   "SDC_EMS01_Carrier74_Faulted" AT %Q10841.6 : Bool;
   "SDC_EMS01_Carrier74_InAuto" AT %Q10841.7 : Bool;
   "SDC_EMS01_Carrier75_Spare0" AT %Q10842.0 : Bool;
   "SDC_EMS01_Carrier75_DriveTripped" AT %Q10842.1 : Bool;
   "SDC_EMS01_Carrier75_Spare2" AT %Q10842.2 : Bool;
   "SDC_EMS01_Carrier75_PositioningComplete" AT %Q10842.3 : Bool;
   "SDC_EMS01_Carrier75_RunStopPressed" AT %Q10842.4 : Bool;
   "SDC_EMS01_Carrier75_Moving" AT %Q10842.5 : Bool;
   "SDC_EMS01_Carrier75_Faulted" AT %Q10842.6 : Bool;
   "SDC_EMS01_Carrier75_InAuto" AT %Q10842.7 : Bool;
   "SDC_EMS01_Carrier76_Spare0" AT %Q10843.0 : Bool;
   "SDC_EMS01_Carrier76_DriveTripped" AT %Q10843.1 : Bool;
   "SDC_EMS01_Carrier76_Spare2" AT %Q10843.2 : Bool;
   "SDC_EMS01_Carrier76_PositioningComplete" AT %Q10843.3 : Bool;
   "SDC_EMS01_Carrier76_RunStopPressed" AT %Q10843.4 : Bool;
   "SDC_EMS01_Carrier76_Moving" AT %Q10843.5 : Bool;
   "SDC_EMS01_Carrier76_Faulted" AT %Q10843.6 : Bool;
   "SDC_EMS01_Carrier76_InAuto" AT %Q10843.7 : Bool;
   "SDC_EMS01_Carrier77_Spare0" AT %Q10844.0 : Bool;
   "SDC_EMS01_Carrier77_DriveTripped" AT %Q10844.1 : Bool;
   "SDC_EMS01_Carrier77_Spare2" AT %Q10844.2 : Bool;
   "SDC_EMS01_Carrier77_PositioningComplete" AT %Q10844.3 : Bool;
   "SDC_EMS01_Carrier77_RunStopPressed" AT %Q10844.4 : Bool;
   "SDC_EMS01_Carrier77_Moving" AT %Q10844.5 : Bool;
   "SDC_EMS01_Carrier77_Faulted" AT %Q10844.6 : Bool;
   "SDC_EMS01_Carrier77_InAuto" AT %Q10844.7 : Bool;
   "SDC_EMS01_Carrier78_Spare0" AT %Q10845.0 : Bool;
   "SDC_EMS01_Carrier78_DriveTripped" AT %Q10845.1 : Bool;
   "SDC_EMS01_Carrier78_Spare2" AT %Q10845.2 : Bool;
   "SDC_EMS01_Carrier78_PositioningComplete" AT %Q10845.3 : Bool;
   "SDC_EMS01_Carrier78_RunStopPressed" AT %Q10845.4 : Bool;
   "SDC_EMS01_Carrier78_Moving" AT %Q10845.5 : Bool;
   "SDC_EMS01_Carrier78_Faulted" AT %Q10845.6 : Bool;
   "SDC_EMS01_Carrier78_InAuto" AT %Q10845.7 : Bool;
   "SDC_EMS01_Carrier79_Spare0" AT %Q10846.0 : Bool;
   "SDC_EMS01_Carrier79_DriveTripped" AT %Q10846.1 : Bool;
   "SDC_EMS01_Carrier79_Spare2" AT %Q10846.2 : Bool;
   "SDC_EMS01_Carrier79_PositioningComplete" AT %Q10846.3 : Bool;
   "SDC_EMS01_Carrier79_RunStopPressed" AT %Q10846.4 : Bool;
   "SDC_EMS01_Carrier79_Moving" AT %Q10846.5 : Bool;
   "SDC_EMS01_Carrier79_Faulted" AT %Q10846.6 : Bool;
   "SDC_EMS01_Carrier79_InAuto" AT %Q10846.7 : Bool;
   "SDC_EMS01_Carrier80_Spare0" AT %Q10847.0 : Bool;
   "SDC_EMS01_Carrier80_DriveTripped" AT %Q10847.1 : Bool;
   "SDC_EMS01_Carrier80_Spare2" AT %Q10847.2 : Bool;
   "SDC_EMS01_Carrier80_PositioningComplete" AT %Q10847.3 : Bool;
   "SDC_EMS01_Carrier80_RunStopPressed" AT %Q10847.4 : Bool;
   "SDC_EMS01_Carrier80_Moving" AT %Q10847.5 : Bool;
   "SDC_EMS01_Carrier80_Faulted" AT %Q10847.6 : Bool;
   "SDC_EMS01_Carrier80_InAuto" AT %Q10847.7 : Bool;
   "SDC_EMS01_Carrier81_Spare0" AT %Q10848.0 : Bool;
   "SDC_EMS01_Carrier81_DriveTripped" AT %Q10848.1 : Bool;
   "SDC_EMS01_Carrier81_Spare2" AT %Q10848.2 : Bool;
   "SDC_EMS01_Carrier81_PositioningComplete" AT %Q10848.3 : Bool;
   "SDC_EMS01_Carrier81_RunStopPressed" AT %Q10848.4 : Bool;
   "SDC_EMS01_Carrier81_Moving" AT %Q10848.5 : Bool;
   "SDC_EMS01_Carrier81_Faulted" AT %Q10848.6 : Bool;
   "SDC_EMS01_Carrier81_InAuto" AT %Q10848.7 : Bool;
   "SDC_EMS01_Carrier82_Spare0" AT %Q10849.0 : Bool;
   "SDC_EMS01_Carrier82_DriveTripped" AT %Q10849.1 : Bool;
   "SDC_EMS01_Carrier82_Spare2" AT %Q10849.2 : Bool;
   "SDC_EMS01_Carrier82_PositioningComplete" AT %Q10849.3 : Bool;
   "SDC_EMS01_Carrier82_RunStopPressed" AT %Q10849.4 : Bool;
   "SDC_EMS01_Carrier82_Moving" AT %Q10849.5 : Bool;
   "SDC_EMS01_Carrier82_Faulted" AT %Q10849.6 : Bool;
   "SDC_EMS01_Carrier82_InAuto" AT %Q10849.7 : Bool;
   "SDC_EMS01_Carrier83_Spare0" AT %Q10850.0 : Bool;
   "SDC_EMS01_Carrier83_DriveTripped" AT %Q10850.1 : Bool;
   "SDC_EMS01_Carrier83_Spare2" AT %Q10850.2 : Bool;
   "SDC_EMS01_Carrier83_PositioningComplete" AT %Q10850.3 : Bool;
   "SDC_EMS01_Carrier83_RunStopPressed" AT %Q10850.4 : Bool;
   "SDC_EMS01_Carrier83_Moving" AT %Q10850.5 : Bool;
   "SDC_EMS01_Carrier83_Faulted" AT %Q10850.6 : Bool;
   "SDC_EMS01_Carrier83_InAuto" AT %Q10850.7 : Bool;
   "SDC_EMS01_Carrier84_Spare0" AT %Q10851.0 : Bool;
   "SDC_EMS01_Carrier84_DriveTripped" AT %Q10851.1 : Bool;
   "SDC_EMS01_Carrier84_Spare2" AT %Q10851.2 : Bool;
   "SDC_EMS01_Carrier84_PositioningComplete" AT %Q10851.3 : Bool;
   "SDC_EMS01_Carrier84_RunStopPressed" AT %Q10851.4 : Bool;
   "SDC_EMS01_Carrier84_Moving" AT %Q10851.5 : Bool;
   "SDC_EMS01_Carrier84_Faulted" AT %Q10851.6 : Bool;
   "SDC_EMS01_Carrier84_InAuto" AT %Q10851.7 : Bool;
   "SDC_EMS01_Carrier85_Spare0" AT %Q10852.0 : Bool;
   "SDC_EMS01_Carrier85_DriveTripped" AT %Q10852.1 : Bool;
   "SDC_EMS01_Carrier85_Spare2" AT %Q10852.2 : Bool;
   "SDC_EMS01_Carrier85_PositioningComplete" AT %Q10852.3 : Bool;
   "SDC_EMS01_Carrier85_RunStopPressed" AT %Q10852.4 : Bool;
   "SDC_EMS01_Carrier85_Moving" AT %Q10852.5 : Bool;
   "SDC_EMS01_Carrier85_Faulted" AT %Q10852.6 : Bool;
   "SDC_EMS01_Carrier85_InAuto" AT %Q10852.7 : Bool;
   "SDC_EMS01_Carrier86_Spare0" AT %Q10853.0 : Bool;
   "SDC_EMS01_Carrier86_DriveTripped" AT %Q10853.1 : Bool;
   "SDC_EMS01_Carrier86_Spare2" AT %Q10853.2 : Bool;
   "SDC_EMS01_Carrier86_PositioningComplete" AT %Q10853.3 : Bool;
   "SDC_EMS01_Carrier86_RunStopPressed" AT %Q10853.4 : Bool;
   "SDC_EMS01_Carrier86_Moving" AT %Q10853.5 : Bool;
   "SDC_EMS01_Carrier86_Faulted" AT %Q10853.6 : Bool;
   "SDC_EMS01_Carrier86_InAuto" AT %Q10853.7 : Bool;
   "SDC_EMS01_Carrier87_Spare0" AT %Q10854.0 : Bool;
   "SDC_EMS01_Carrier87_DriveTripped" AT %Q10854.1 : Bool;
   "SDC_EMS01_Carrier87_Spare2" AT %Q10854.2 : Bool;
   "SDC_EMS01_Carrier87_PositioningComplete" AT %Q10854.3 : Bool;
   "SDC_EMS01_Carrier87_RunStopPressed" AT %Q10854.4 : Bool;
   "SDC_EMS01_Carrier87_Moving" AT %Q10854.5 : Bool;
   "SDC_EMS01_Carrier87_Faulted" AT %Q10854.6 : Bool;
   "SDC_EMS01_Carrier87_InAuto" AT %Q10854.7 : Bool;
   "SDC_EMS01_Carrier88_Spare0" AT %Q10855.0 : Bool;
   "SDC_EMS01_Carrier88_DriveTripped" AT %Q10855.1 : Bool;
   "SDC_EMS01_Carrier88_Spare2" AT %Q10855.2 : Bool;
   "SDC_EMS01_Carrier88_PositioningComplete" AT %Q10855.3 : Bool;
   "SDC_EMS01_Carrier88_RunStopPressed" AT %Q10855.4 : Bool;
   "SDC_EMS01_Carrier88_Moving" AT %Q10855.5 : Bool;
   "SDC_EMS01_Carrier88_Faulted" AT %Q10855.6 : Bool;
   "SDC_EMS01_Carrier88_InAuto" AT %Q10855.7 : Bool;
   "SDC_EMS01_Carrier89_Spare0" AT %Q10856.0 : Bool;
   "SDC_EMS01_Carrier89_DriveTripped" AT %Q10856.1 : Bool;
   "SDC_EMS01_Carrier89_Spare2" AT %Q10856.2 : Bool;
   "SDC_EMS01_Carrier89_PositioningComplete" AT %Q10856.3 : Bool;
   "SDC_EMS01_Carrier89_RunStopPressed" AT %Q10856.4 : Bool;
   "SDC_EMS01_Carrier89_Moving" AT %Q10856.5 : Bool;
   "SDC_EMS01_Carrier89_Faulted" AT %Q10856.6 : Bool;
   "SDC_EMS01_Carrier89_InAuto" AT %Q10856.7 : Bool;
   "SDC_EMS01_Carrier90_Spare0" AT %Q10857.0 : Bool;
   "SDC_EMS01_Carrier90_DriveTripped" AT %Q10857.1 : Bool;
   "SDC_EMS01_Carrier90_Spare2" AT %Q10857.2 : Bool;
   "SDC_EMS01_Carrier90_PositioningComplete" AT %Q10857.3 : Bool;
   "SDC_EMS01_Carrier90_RunStopPressed" AT %Q10857.4 : Bool;
   "SDC_EMS01_Carrier90_Moving" AT %Q10857.5 : Bool;
   "SDC_EMS01_Carrier90_Faulted" AT %Q10857.6 : Bool;
   "SDC_EMS01_Carrier90_InAuto" AT %Q10857.7 : Bool;
   "SDC_EMS01_Carrier91_Spare0" AT %Q10858.0 : Bool;
   "SDC_EMS01_Carrier91_DriveTripped" AT %Q10858.1 : Bool;
   "SDC_EMS01_Carrier91_Spare2" AT %Q10858.2 : Bool;
   "SDC_EMS01_Carrier91_PositioningComplete" AT %Q10858.3 : Bool;
   "SDC_EMS01_Carrier91_RunStopPressed" AT %Q10858.4 : Bool;
   "SDC_EMS01_Carrier91_Moving" AT %Q10858.5 : Bool;
   "SDC_EMS01_Carrier91_Faulted" AT %Q10858.6 : Bool;
   "SDC_EMS01_Carrier91_InAuto" AT %Q10858.7 : Bool;
   "SDC_EMS01_Carrier92_Spare0" AT %Q10859.0 : Bool;
   "SDC_EMS01_Carrier92_DriveTripped" AT %Q10859.1 : Bool;
   "SDC_EMS01_Carrier92_Spare2" AT %Q10859.2 : Bool;
   "SDC_EMS01_Carrier92_PositioningComplete" AT %Q10859.3 : Bool;
   "SDC_EMS01_Carrier92_RunStopPressed" AT %Q10859.4 : Bool;
   "SDC_EMS01_Carrier92_Moving" AT %Q10859.5 : Bool;
   "SDC_EMS01_Carrier92_Faulted" AT %Q10859.6 : Bool;
   "SDC_EMS01_Carrier92_InAuto" AT %Q10859.7 : Bool;
   "SDC_EMS01_Carrier93_Spare0" AT %Q10860.0 : Bool;
   "SDC_EMS01_Carrier93_DriveTripped" AT %Q10860.1 : Bool;
   "SDC_EMS01_Carrier93_Spare2" AT %Q10860.2 : Bool;
   "SDC_EMS01_Carrier93_PositioningComplete" AT %Q10860.3 : Bool;
   "SDC_EMS01_Carrier93_RunStopPressed" AT %Q10860.4 : Bool;
   "SDC_EMS01_Carrier93_Moving" AT %Q10860.5 : Bool;
   "SDC_EMS01_Carrier93_Faulted" AT %Q10860.6 : Bool;
   "SDC_EMS01_Carrier93_InAuto" AT %Q10860.7 : Bool;
   "SDC_EMS01_Carrier94_Spare0" AT %Q10861.0 : Bool;
   "SDC_EMS01_Carrier94_DriveTripped" AT %Q10861.1 : Bool;
   "SDC_EMS01_Carrier94_Spare2" AT %Q10861.2 : Bool;
   "SDC_EMS01_Carrier94_PositioningComplete" AT %Q10861.3 : Bool;
   "SDC_EMS01_Carrier94_RunStopPressed" AT %Q10861.4 : Bool;
   "SDC_EMS01_Carrier94_Moving" AT %Q10861.5 : Bool;
   "SDC_EMS01_Carrier94_Faulted" AT %Q10861.6 : Bool;
   "SDC_EMS01_Carrier94_InAuto" AT %Q10861.7 : Bool;
   "SDC_EMS01_Carrier95_Spare0" AT %Q10862.0 : Bool;
   "SDC_EMS01_Carrier95_DriveTripped" AT %Q10862.1 : Bool;
   "SDC_EMS01_Carrier95_Spare2" AT %Q10862.2 : Bool;
   "SDC_EMS01_Carrier95_PositioningComplete" AT %Q10862.3 : Bool;
   "SDC_EMS01_Carrier95_RunStopPressed" AT %Q10862.4 : Bool;
   "SDC_EMS01_Carrier95_Moving" AT %Q10862.5 : Bool;
   "SDC_EMS01_Carrier95_Faulted" AT %Q10862.6 : Bool;
   "SDC_EMS01_Carrier95_InAuto" AT %Q10862.7 : Bool;
   "SDC_EMS01_Carrier1_Fault" AT %QB10512 : Byte;
   "SDC_EMS01_Carrier2_Fault" AT %QB10513 : Byte;
   "SDC_EMS01_Carrier3_Fault" AT %QB10514 : Byte;
   "SDC_EMS01_Carrier4_Fault" AT %QB10515 : Byte;
   "SDC_EMS01_Carrier5_Fault" AT %QB10516 : Byte;
   "SDC_EMS01_Carrier6_Fault" AT %QB10517 : Byte;
   "SDC_EMS01_Carrier7_Fault" AT %QB10518 : Byte;
   "SDC_EMS01_Carrier8_Fault" AT %QB10519 : Byte;
   "SDC_EMS01_Carrier9_Fault" AT %QB10520 : Byte;
   "SDC_EMS01_Carrier10_Fault" AT %QB10521 : Byte;
   "SDC_EMS01_Carrier11_Fault" AT %QB10522 : Byte;
   "SDC_EMS01_Carrier12_Fault" AT %QB10523 : Byte;
   "SDC_EMS01_Carrier13_Fault" AT %QB10524 : Byte;
   "SDC_EMS01_Carrier14_Fault" AT %QB10525 : Byte;
   "SDC_EMS01_Carrier15_Fault" AT %QB10526 : Byte;
   "SDC_EMS01_Carrier16_Fault" AT %QB10527 : Byte;
   "SDC_EMS01_Carrier17_Fault" AT %QB10528 : Byte;
   "SDC_EMS01_Carrier18_Fault" AT %QB10529 : Byte;
   "SDC_EMS01_Carrier19_Fault" AT %QB10530 : Byte;
   "SDC_EMS01_Carrier20_Fault" AT %QB10531 : Byte;
   "SDC_EMS01_Carrier21_Fault" AT %QB10532 : Byte;
   "SDC_EMS01_Carrier22_Fault" AT %QB10533 : Byte;
   "SDC_EMS01_Carrier23_Fault" AT %QB10534 : Byte;
   "SDC_EMS01_Carrier24_Fault" AT %QB10535 : Byte;
   "SDC_EMS01_Carrier25_Fault" AT %QB10536 : Byte;
   "SDC_EMS01_Carrier26_Fault" AT %QB10537 : Byte;
   "SDC_EMS01_Carrier27_Fault" AT %QB10538 : Byte;
   "SDC_EMS01_Carrier28_Fault" AT %QB10539 : Byte;
   "SDC_EMS01_Carrier29_Fault" AT %QB10540 : Byte;
   "SDC_EMS01_Carrier30_Fault" AT %QB10541 : Byte;
   "SDC_EMS01_Carrier31_Fault" AT %QB10542 : Byte;
   "SDC_EMS01_Carrier32_Fault" AT %QB10543 : Byte;
   "SDC_EMS01_Carrier33_Fault" AT %QB10544 : Byte;
   "SDC_EMS01_Carrier34_Fault" AT %QB10545 : Byte;
   "SDC_EMS01_Carrier35_Fault" AT %QB10546 : Byte;
   "SDC_EMS01_Carrier36_Fault" AT %QB10547 : Byte;
   "SDC_EMS01_Carrier37_Fault" AT %QB10548 : Byte;
   "SDC_EMS01_Carrier38_Fault" AT %QB10549 : Byte;
   "SDC_EMS01_Carrier39_Fault" AT %QB10550 : Byte;
   "SDC_EMS01_Carrier40_Fault" AT %QB10551 : Byte;
   "SDC_EMS01_Carrier41_Fault" AT %QB10552 : Byte;
   "SDC_EMS01_Carrier42_Fault" AT %QB10553 : Byte;
   "SDC_EMS01_Carrier43_Fault" AT %QB10554 : Byte;
   "SDC_EMS01_Carrier44_Fault" AT %QB10555 : Byte;
   "SDC_EMS01_Carrier45_Fault" AT %QB10556 : Byte;
   "SDC_EMS01_Carrier46_Fault" AT %QB10557 : Byte;
   "SDC_EMS01_Carrier47_Fault" AT %QB10558 : Byte;
   "SDC_EMS01_Carrier48_Fault" AT %QB10559 : Byte;
   "SDC_EMS01_Carrier49_Fault" AT %QB10560 : Byte;
   "SDC_EMS01_Carrier50_Fault" AT %QB10561 : Byte;
   "SDC_EMS01_Carrier51_Fault" AT %QB10562 : Byte;
   "SDC_EMS01_Carrier52_Fault" AT %QB10563 : Byte;
   "SDC_EMS01_Carrier53_Fault" AT %QB10564 : Byte;
   "SDC_EMS01_Carrier54_Fault" AT %QB10565 : Byte;
   "SDC_EMS01_Carrier55_Fault" AT %QB10566 : Byte;
   "SDC_EMS01_Carrier56_Fault" AT %QB10567 : Byte;
   "SDC_EMS01_Carrier57_Fault" AT %QB10568 : Byte;
   "SDC_EMS01_Carrier58_Fault" AT %QB10569 : Byte;
   "SDC_EMS01_Carrier59_Fault" AT %QB10570 : Byte;
   "SDC_EMS01_Carrier60_Fault" AT %QB10571 : Byte;
   "SDC_EMS01_Carrier61_Fault" AT %QB10572 : Byte;
   "SDC_EMS01_Carrier62_Fault" AT %QB10573 : Byte;
   "SDC_EMS01_Carrier63_Fault" AT %QB10574 : Byte;
   "SDC_EMS01_Carrier64_Fault" AT %QB10575 : Byte;
   "SDC_EMS01_Carrier65_Fault" AT %QB10576 : Byte;
   "SDC_EMS01_Carrier66_Fault" AT %QB10577 : Byte;
   "SDC_EMS01_Carrier67_Fault" AT %QB10578 : Byte;
   "SDC_EMS01_Carrier68_Fault" AT %QB10579 : Byte;
   "SDC_EMS01_Carrier69_Fault" AT %QB10580 : Byte;
   "SDC_EMS01_Carrier70_Fault" AT %QB10581 : Byte;
   "SDC_EMS01_Carrier71_Fault" AT %QB10582 : Byte;
   "SDC_EMS01_Carrier72_Fault" AT %QB10583 : Byte;
   "SDC_EMS01_Carrier73_Fault" AT %QB10584 : Byte;
   "SDC_EMS01_Carrier74_Fault" AT %QB10585 : Byte;
   "SDC_EMS01_Carrier75_Fault" AT %QB10586 : Byte;
   "SDC_EMS01_Carrier76_Fault" AT %QB10587 : Byte;
   "SDC_EMS01_Carrier77_Fault" AT %QB10588 : Byte;
   "SDC_EMS01_Carrier78_Fault" AT %QB10589 : Byte;
   "SDC_EMS01_Carrier79_Fault" AT %QB10590 : Byte;
   "SDC_EMS01_Carrier80_Fault" AT %QB10591 : Byte;
   "SDC_EMS01_Carrier81_Fault" AT %QB10592 : Byte;
   "SDC_EMS01_Carrier82_Fault" AT %QB10593 : Byte;
   "SDC_EMS01_Carrier1_Status" AT %QB10768 : Byte;
   "SDC_EMS01_Carrier2_Status" AT %QB10769 : Byte;
   "SDC_EMS01_Carrier3_Status" AT %QB10770 : Byte;
   "SDC_EMS01_Carrier4_Status" AT %QB10771 : Byte;
   "SDC_EMS01_Carrier5_Status" AT %QB10772 : Byte;
   "SDC_EMS01_Carrier6_Status" AT %QB10773 : Byte;
   "SDC_EMS01_Carrier7_Status" AT %QB10774 : Byte;
   "SDC_EMS01_Carrier8_Status" AT %QB10775 : Byte;
   "SDC_EMS01_Carrier9_Status" AT %QB10776 : Byte;
   "SDC_EMS01_Carrier10_Status" AT %QB10777 : Byte;
   "SDC_EMS01_Carrier11_Status" AT %QB10778 : Byte;
   "SDC_EMS01_Carrier12_Status" AT %QB10779 : Byte;
   "SDC_EMS01_Carrier13_Status" AT %QB10780 : Byte;
   "SDC_EMS01_Carrier14_Status" AT %QB10781 : Byte;
   "SDC_EMS01_Carrier15_Status" AT %QB10782 : Byte;
   "SDC_EMS01_Carrier16_Status" AT %QB10783 : Byte;
   "SDC_EMS01_Carrier17_Status" AT %QB10784 : Byte;
   "SDC_EMS01_Carrier18_Status" AT %QB10785 : Byte;
   "SDC_EMS01_Carrier19_Status" AT %QB10786 : Byte;
   "SDC_EMS01_Carrier20_Status" AT %QB10787 : Byte;
   "SDC_EMS01_Carrier21_Status" AT %QB10788 : Byte;
   "SDC_EMS01_Carrier22_Status" AT %QB10789 : Byte;
   "SDC_EMS01_Carrier23_Status" AT %QB10790 : Byte;
   "SDC_EMS01_Carrier24_Status" AT %QB10791 : Byte;
   "SDC_EMS01_Carrier25_Status" AT %QB10792 : Byte;
   "SDC_EMS01_Carrier26_Status" AT %QB10793 : Byte;
   "SDC_EMS01_Carrier27_Status" AT %QB10794 : Byte;
   "SDC_EMS01_Carrier28_Status" AT %QB10795 : Byte;
   "SDC_EMS01_Carrier29_Status" AT %QB10796 : Byte;
   "SDC_EMS01_Carrier30_Status" AT %QB10797 : Byte;
   "SDC_EMS01_Carrier31_Status" AT %QB10798 : Byte;
   "SDC_EMS01_Carrier32_Status" AT %QB10799 : Byte;
   "SDC_EMS01_Carrier33_Status" AT %QB10800 : Byte;
   "SDC_EMS01_Carrier34_Status" AT %QB10801 : Byte;
   "SDC_EMS01_Carrier35_Status" AT %QB10802 : Byte;
   "SDC_EMS01_Carrier36_Status" AT %QB10803 : Byte;
   "SDC_EMS01_Carrier37_Status" AT %QB10804 : Byte;
   "SDC_EMS01_Carrier38_Status" AT %QB10805 : Byte;
   "SDC_EMS01_Carrier39_Status" AT %QB10806 : Byte;
   "SDC_EMS01_Carrier40_Status" AT %QB10807 : Byte;
   "SDC_EMS01_Carrier41_Status" AT %QB10808 : Byte;
   "SDC_EMS01_Carrier42_Status" AT %QB10809 : Byte;
   "SDC_EMS01_Carrier43_Status" AT %QB10810 : Byte;
   "SDC_EMS01_Carrier44_Status" AT %QB10811 : Byte;
   "SDC_EMS01_Carrier45_Status" AT %QB10812 : Byte;
   "SDC_EMS01_Carrier46_Status" AT %QB10813 : Byte;
   "SDC_EMS01_Carrier47_Status" AT %QB10814 : Byte;
   "SDC_EMS01_Carrier48_Status" AT %QB10815 : Byte;
   "SDC_EMS01_Carrier49_Status" AT %QB10816 : Byte;
   "SDC_EMS01_Carrier50_Status" AT %QB10817 : Byte;
   "SDC_EMS01_Carrier51_Status" AT %QB10818 : Byte;
   "SDC_EMS01_Carrier52_Status" AT %QB10819 : Byte;
   "SDC_EMS01_Carrier53_Status" AT %QB10820 : Byte;
   "SDC_EMS01_Carrier54_Status" AT %QB10821 : Byte;
   "SDC_EMS01_Carrier55_Status" AT %QB10822 : Byte;
   "SDC_EMS01_Carrier56_Status" AT %QB10823 : Byte;
   "SDC_EMS01_Carrier57_Status" AT %QB10824 : Byte;
   "SDC_EMS01_Carrier58_Status" AT %QB10825 : Byte;
   "SDC_EMS01_Carrier59_Status" AT %QB10826 : Byte;
   "SDC_EMS01_Carrier60_Status" AT %QB10827 : Byte;
   "SDC_EMS01_Carrier61_Status" AT %QB10828 : Byte;
   "SDC_EMS01_Carrier62_Status" AT %QB10829 : Byte;
   "SDC_EMS01_Carrier63_Status" AT %QB10830 : Byte;
   "SDC_EMS01_Carrier64_Status" AT %QB10831 : Byte;
   "SDC_EMS01_Carrier65_Status" AT %QB10832 : Byte;
   "SDC_EMS01_Carrier66_Status" AT %QB10833 : Byte;
   "SDC_EMS01_Carrier67_Status" AT %QB10834 : Byte;
   "SDC_EMS01_Carrier68_Status" AT %QB10835 : Byte;
   "SDC_EMS01_Carrier69_Status" AT %QB10836 : Byte;
   "SDC_EMS01_Carrier70_Status" AT %QB10837 : Byte;
   "SDC_EMS01_Carrier71_Status" AT %QB10838 : Byte;
   "SDC_EMS01_Carrier72_Status" AT %QB10839 : Byte;
   "SDC_EMS01_Carrier73_Status" AT %QB10840 : Byte;
   "SDC_EMS01_Carrier74_Status" AT %QB10841 : Byte;
   "SDC_EMS01_Carrier75_Status" AT %QB10842 : Byte;
   "SDC_EMS01_Carrier76_Status" AT %QB10843 : Byte;
   "SDC_EMS01_Carrier77_Status" AT %QB10844 : Byte;
   "SDC_EMS01_Carrier78_Status" AT %QB10845 : Byte;
   "SDC_EMS01_Carrier79_Status" AT %QB10846 : Byte;
   "SDC_EMS01_Carrier80_Status" AT %QB10847 : Byte;
   "SDC_EMS01_Carrier81_Status" AT %QB10848 : Byte;
   "SDC_EMS01_Carrier82_Status" AT %QB10849 : Byte;
   "SDC_EMS01_Carrier83_Status" AT %QB10850 : Byte;
   "SDC_EMS01_Carrier84_Status" AT %QB10851 : Byte;
   "SDC_EMS01_Carrier85_Status" AT %QB10852 : Byte;
   "SDC_EMS01_Carrier86_Status" AT %QB10853 : Byte;
   "SDC_EMS01_Carrier87_Status" AT %QB10854 : Byte;
   "SDC_EMS01_Carrier88_Status" AT %QB10855 : Byte;
   "SDC_EMS01_Carrier89_Status" AT %QB10856 : Byte;
   "SDC_EMS01_Carrier90_Status" AT %QB10857 : Byte;
   "SDC_EMS01_Carrier91_Status" AT %QB10858 : Byte;
   "SDC_EMS01_Carrier92_Status" AT %QB10859 : Byte;
   "SDC_EMS01_Carrier93_Status" AT %QB10860 : Byte;
   "SDC_EMS01_Carrier94_Status" AT %QB10861 : Byte;
   "SDC_EMS01_Carrier95_Status" AT %QB10862 : Byte;
   "SDC_EMS01_Carrier1_Zone" AT %QB10328 : Byte;
   "SDC_EMS01_Carrier2_Zone" AT %QB10329 : Byte;
   "SDC_EMS01_Carrier3_Zone" AT %QB10330 : Byte;
   "SDC_EMS01_Carrier4_Zone" AT %QB10331 : Byte;
   "SDC_EMS01_Carrier5_Zone" AT %QB10332 : Byte;
   "SDC_EMS01_Carrier6_Zone" AT %QB10333 : Byte;
   "SDC_EMS01_Carrier7_Zone" AT %QB10334 : Byte;
   "SDC_EMS01_Carrier8_Zone" AT %QB10335 : Byte;
   "SDC_EMS01_Carrier9_Zone" AT %QB10336 : Byte;
   "SDC_EMS01_Carrier10_Zone" AT %QB10337 : Byte;
   "SDC_EMS01_Carrier11_Zone" AT %QB10338 : Byte;
   "SDC_EMS01_Carrier12_Zone" AT %QB10339 : Byte;
   "SDC_EMS01_Carrier13_Zone" AT %QB10340 : Byte;
   "SDC_EMS01_Carrier14_Zone" AT %QB10341 : Byte;
   "SDC_EMS01_Carrier15_Zone" AT %QB10342 : Byte;
   "SDC_EMS01_Carrier16_Zone" AT %QB10343 : Byte;
   "SDC_EMS01_Carrier17_Zone" AT %QB10344 : Byte;
   "SDC_EMS01_Carrier18_Zone" AT %QB10345 : Byte;
   "SDC_EMS01_Carrier19_Zone" AT %QB10346 : Byte;
   "SDC_EMS01_Carrier20_Zone" AT %QB10347 : Byte;
   "SDC_EMS01_Carrier21_Zone" AT %QB10348 : Byte;
   "SDC_EMS01_Carrier22_Zone" AT %QB10349 : Byte;
   "SDC_EMS01_Carrier23_Zone" AT %QB10350 : Byte;
   "SDC_EMS01_Carrier24_Zone" AT %QB10351 : Byte;
   "SDC_EMS01_Carrier25_Zone" AT %QB10352 : Byte;
   "SDC_EMS01_Carrier26_Zone" AT %QB10353 : Byte;
   "SDC_EMS01_Carrier27_Zone" AT %QB10354 : Byte;
   "SDC_EMS01_Carrier28_Zone" AT %QB10355 : Byte;
   "SDC_EMS01_Carrier29_Zone" AT %QB10356 : Byte;
   "SDC_EMS01_Carrier30_Zone" AT %QB10357 : Byte;
   "SDC_EMS01_Carrier31_Zone" AT %QB10358 : Byte;
   "SDC_EMS01_Carrier32_Zone" AT %QB10359 : Byte;
   "SDC_EMS01_Carrier33_Zone" AT %QB10360 : Byte;
   "SDC_EMS01_Carrier34_Zone" AT %QB10361 : Byte;
   "SDC_EMS01_Carrier35_Zone" AT %QB10362 : Byte;
   "SDC_EMS01_Carrier36_Zone" AT %QB10363 : Byte;
   "SDC_EMS01_Carrier37_Zone" AT %QB10364 : Byte;
   "SDC_EMS01_Carrier38_Zone" AT %QB10365 : Byte;
   "SDC_EMS01_Carrier39_Zone" AT %QB10366 : Byte;
   "SDC_EMS01_Carrier40_Zone" AT %QB10367 : Byte;
   "SDC_EMS01_Carrier41_Zone" AT %QB10368 : Byte;
   "SDC_EMS01_Carrier42_Zone" AT %QB10369 : Byte;
   "SDC_EMS01_Carrier43_Zone" AT %QB10370 : Byte;
   "SDC_EMS01_Carrier44_Zone" AT %QB10371 : Byte;
   "SDC_EMS01_Carrier45_Zone" AT %QB10372 : Byte;
   "SDC_EMS01_Carrier46_Zone" AT %QB10373 : Byte;
   "SDC_EMS01_Carrier47_Zone" AT %QB10374 : Byte;
   "SDC_EMS01_Carrier48_Zone" AT %QB10375 : Byte;
   "SDC_EMS01_Carrier49_Zone" AT %QB10376 : Byte;
   "SDC_EMS01_Carrier50_Zone" AT %QB10377 : Byte;
   "SDC_EMS01_Carrier51_Zone" AT %QB10378 : Byte;
   "SDC_EMS01_Carrier52_Zone" AT %QB10379 : Byte;
   "SDC_EMS01_Carrier53_Zone" AT %QB10380 : Byte;
   "SDC_EMS01_Carrier54_Zone" AT %QB10381 : Byte;
   "SDC_EMS01_Carrier55_Zone" AT %QB10382 : Byte;
   "SDC_EMS01_Carrier56_Zone" AT %QB10383 : Byte;
   "SDC_EMS01_Carrier57_Zone" AT %QB10384 : Byte;
   "SDC_EMS01_Carrier58_Zone" AT %QB10385 : Byte;
   "SDC_EMS01_Carrier59_Zone" AT %QB10386 : Byte;
   "SDC_EMS01_Carrier60_Zone" AT %QB10387 : Byte;
   "SDC_EMS01_Carrier61_Zone" AT %QB10388 : Byte;
   "SDC_EMS01_Carrier62_Zone" AT %QB10389 : Byte;
   "SDC_EMS01_Carrier63_Zone" AT %QB10390 : Byte;
   "SDC_EMS01_Carrier64_Zone" AT %QB10391 : Byte;
   "SDC_EMS01_Carrier65_Zone" AT %QB10392 : Byte;
   "SDC_EMS01_Carrier66_Zone" AT %QB10393 : Byte;
   "SDC_EMS01_Carrier67_Zone" AT %QB10394 : Byte;
   "SDC_EMS01_Carrier68_Zone" AT %QB10395 : Byte;
   "SDC_EMS01_Carrier69_Zone" AT %QB10396 : Byte;
   "SDC_EMS01_Carrier70_Zone" AT %QB10397 : Byte;
   "SDC_EMS01_Carrier71_Zone" AT %QB10398 : Byte;
   "SDC_EMS01_Carrier72_Zone" AT %QB10399 : Byte;
   "SDC_EMS01_Carrier73_Zone" AT %QB10400 : Byte;
   "SDC_EMS01_Carrier74_Zone" AT %QB10401 : Byte;
   "SDC_EMS01_Carrier75_Zone" AT %QB10402 : Byte;
   "SDC_EMS01_Carrier76_Zone" AT %QB10403 : Byte;
   "SDC_EMS01_Carrier77_Zone" AT %QB10404 : Byte;
   "SDC_EMS01_Carrier78_Zone" AT %QB10405 : Byte;
   "SDC_EMS01_Carrier79_Zone" AT %QB10406 : Byte;
   "SDC_EMS01_Carrier80_Zone" AT %QB10407 : Byte;
   "SDC_EMS01_Carrier81_Zone" AT %QB10408 : Byte;
   "SDC_EMS01_Carrier82_Zone" AT %QB10409 : Byte;
   "SDC_EMS01_Stop1_Status" AT %QW11024 : Word;
   "SDC_EMS01_Stop2_Status" AT %QW11026 : Word;
   "SDC_EMS01_Stop3_Status" AT %QW11028 : Word;
   "SDC_EMS01_Stop4_Status" AT %QW11030 : Word;
   "SDC_EMS01_Stop5_Status" AT %QW11032 : Word;
   "SDC_EMS01_Stop6_Status" AT %QW11034 : Word;
   "SDC_EMS01_Stop7_Status" AT %QW11036 : Word;
   "SDC_EMS01_Stop8_Status" AT %QW11038 : Word;
   "SDC_EMS01_Stop9_Status" AT %QW11040 : Word;
   "SDC_EMS01_Stop10_Status" AT %QW11042 : Word;
   "SDC_EMS01_Stop11_Status" AT %QW11044 : Word;
   "SDC_EMS01_Stop12_Status" AT %QW11046 : Word;
   "SDC_EMS01_Stop13_Status" AT %QW11048 : Word;
   "SDC_EMS01_Stop14_Status" AT %QW11050 : Word;
   "SDC_EMS01_Stop15_Status" AT %QW11052 : Word;
   "SDC_EMS01_Stop16_Status" AT %QW11054 : Word;
   "SDC_EMS01_Stop17_Status" AT %QW11056 : Word;
   "SDC_EMS01_Stop18_Status" AT %QW11058 : Word;
   "SDC_EMS01_Stop19_Status" AT %QW11060 : Word;
   "SDC_EMS01_Stop20_Status" AT %QW11062 : Word;
   "SDC_EMS01_Stop21_Status" AT %QW11064 : Word;
   "SDC_EMS01_Stop22_Status" AT %QW11066 : Word;
   "SDC_EMS01_Stop23_Status" AT %QW11068 : Word;
   "SDC_EMS01_Stop24_Status" AT %QW11070 : Word;
   "SDC_EMS01_Stop25_Status" AT %QW11072 : Word;
   "SDC_EMS01_Stop26_Status" AT %QW11074 : Word;
   "SDC_EMS01_Stop27_Status" AT %QW11076 : Word;
   "SDC_EMS01_Stop28_Status" AT %QW11078 : Word;
   "SDC_EMS01_Stop29_Status" AT %QW11080 : Word;
   "SDC_EMS01_Stop30_Status" AT %QW11082 : Word;
   "SDC_EMS01_Stop31_Status" AT %QW11084 : Word;
   "SDC_EMS01_Stop32_Status" AT %QW11086 : Word;
   "SDC_EMS01_Stop33_Status" AT %QW11088 : Word;
   "SDC_EMS01_Stop34_Status" AT %QW11090 : Word;
   "SDC_EMS01_Stop35_Status" AT %QW11092 : Word;
   "SDC_EMS01_Stop36_Status" AT %QW11094 : Word;
   "SDC_EMS01_Stop37_Status" AT %QW11096 : Word;
   "SDC_EMS01_Stop38_Status" AT %QW11098 : Word;
   "SDC_EMS01_Stop39_Status" AT %QW11100 : Word;
   "SDC_EMS01_Stop40_Status" AT %QW11102 : Word;
   "SDC_EMS01_Stop41_Status" AT %QW11104 : Word;
   "SDC_EMS01_Stop42_Status" AT %QW11106 : Word;
   "SDC_EMS01_Stop43_Status" AT %QW11108 : Word;
   "SDC_EMS01_Stop44_Status" AT %QW11110 : Word;
   "SDC_EMS01_Stop45_Status" AT %QW11112 : Word;
   "SDC_EMS01_Stop46_Status" AT %QW11114 : Word;
   "SDC_EMS01_Stop47_Status" AT %QW11116 : Word;
   "SDC_EMS01_Stop48_Status" AT %QW11118 : Word;
   "SDC_EMS01_Stop49_Status" AT %QW11120 : Word;
   "SDC_EMS01_Stop50_Status" AT %QW11122 : Word;
   "SDC_EMS01_Stop51_Status" AT %QW11124 : Word;
   "SDC_EMS01_Stop52_Status" AT %QW11126 : Word;
   "SDC_EMS01_Stop53_Status" AT %QW11128 : Word;
   "SDC_EMS01_Stop54_Status" AT %QW11130 : Word;
   "SDC_EMS01_Stop55_Status" AT %QW11132 : Word;
   "SDC_EMS01_Stop56_Status" AT %QW11134 : Word;
   "SDC_EMS01_Stop57_Status" AT %QW11136 : Word;
   "SDC_EMS01_Stop58_Status" AT %QW11138 : Word;
   "SDC_EMS01_Stop59_Status" AT %QW11140 : Word;
   "SDC_EMS01_Stop60_Status" AT %QW11142 : Word;
   "SDC_EMS01_Stop61_Status" AT %QW11144 : Word;
   "SDC_EMS01_Stop62_Status" AT %QW11146 : Word;
   "SDC_EMS01_Stop63_Status" AT %QW11148 : Word;
   "SDC_EMS01_Stop64_Status" AT %QW11150 : Word;
   "SDC_EMS01_Stop65_Status" AT %QW11152 : Word;
   "SDC_EMS01_Carrier1_Position" AT %QD10000 : DWord;
   "SDC_EMS01_Carrier2_Position" AT %QD10004 : DWord;
   "SDC_EMS01_Carrier3_Position" AT %QD10008 : DWord;
   "SDC_EMS01_Carrier4_Position" AT %QD10012 : DWord;
   "SDC_EMS01_Carrier5_Position" AT %QD10016 : DWord;
   "SDC_EMS01_Carrier6_Position" AT %QD10020 : DWord;
   "SDC_EMS01_Carrier7_Position" AT %QD10024 : DWord;
   "SDC_EMS01_Carrier8_Position" AT %QD10028 : DWord;
   "SDC_EMS01_Carrier9_Position" AT %QD10032 : DWord;
   "SDC_EMS01_Carrier10_Position" AT %QD10036 : DWord;
   "SDC_EMS01_Carrier11_Position" AT %QD10040 : DWord;
   "SDC_EMS01_Carrier12_Position" AT %QD10044 : DWord;
   "SDC_EMS01_Carrier13_Position" AT %QD10048 : DWord;
   "SDC_EMS01_Carrier14_Position" AT %QD10052 : DWord;
   "SDC_EMS01_Carrier15_Position" AT %QD10056 : DWord;
   "SDC_EMS01_Carrier16_Position" AT %QD10060 : DWord;
   "SDC_EMS01_Carrier17_Position" AT %QD10064 : DWord;
   "SDC_EMS01_Carrier18_Position" AT %QD10068 : DWord;
   "SDC_EMS01_Carrier19_Position" AT %QD10072 : DWord;
   "SDC_EMS01_Carrier20_Position" AT %QD10076 : DWord;
   "SDC_EMS01_Carrier21_Position" AT %QD10080 : DWord;
   "SDC_EMS01_Carrier22_Position" AT %QD10084 : DWord;
   "SDC_EMS01_Carrier23_Position" AT %QD10088 : DWord;
   "SDC_EMS01_Carrier24_Position" AT %QD10092 : DWord;
   "SDC_EMS01_Carrier25_Position" AT %QD10096 : DWord;
   "SDC_EMS01_Carrier28_Position" AT %QD10108 : DWord;
   "SDC_EMS01_Carrier29_Position" AT %QD10112 : DWord;
   "SDC_EMS01_Carrier30_Position" AT %QD10116 : DWord;
   "SDC_EMS01_Carrier31_Position" AT %QD10120 : DWord;
   "SDC_EMS01_Carrier32_Position" AT %QD10124 : DWord;
   "SDC_EMS01_Carrier33_Position" AT %QD10128 : DWord;
   "SDC_EMS01_Carrier34_Position" AT %QD10132 : DWord;
   "SDC_EMS01_Carrier35_Position" AT %QD10136 : DWord;
   "SDC_EMS01_Carrier36_Position" AT %QD10140 : DWord;
   "SDC_EMS01_Carrier37_Position" AT %QD10144 : DWord;
   "SDC_EMS01_Carrier38_Position" AT %QD10148 : DWord;
   "SDC_EMS01_Carrier39_Position" AT %QD10152 : DWord;
   "SDC_EMS01_Carrier40_Position" AT %QD10156 : DWord;
   "SDC_EMS01_Carrier41_Position" AT %QD10160 : DWord;
   "SDC_EMS01_Carrier42_Position" AT %QD10164 : DWord;
   "SDC_EMS01_Carrier43_Position" AT %QD10168 : DWord;
   "SDC_EMS01_Carrier44_Position" AT %QD10172 : DWord;
   "SDC_EMS01_Carrier45_Position" AT %QD10176 : DWord;
   "SDC_EMS01_Carrier46_Position" AT %QD10180 : DWord;
   "SDC_EMS01_Carrier47_Position" AT %QD10184 : DWord;
   "SDC_EMS01_Carrier48_Position" AT %QD10188 : DWord;
   "SDC_EMS01_Carrier49_Position" AT %QD10192 : DWord;
   "SDC_EMS01_Carrier50_Position" AT %QD10196 : DWord;
   "SDC_EMS01_Carrier51_Position" AT %QD10200 : DWord;
   "SDC_EMS01_Carrier52_Position" AT %QD10204 : DWord;
   "SDC_EMS01_Carrier53_Position" AT %QD10208 : DWord;
   "SDC_EMS01_Carrier54_Position" AT %QD10212 : DWord;
   "SDC_EMS01_Carrier55_Position" AT %QD10216 : DWord;
   "SDC_EMS01_Carrier56_Position" AT %QD10220 : DWord;
   "SDC_EMS01_Carrier57_Position" AT %QD10224 : DWord;
   "SDC_EMS01_Carrier58_Position" AT %QD10228 : DWord;
   "SDC_EMS01_Carrier59_Position" AT %QD10232 : DWord;
   "SDC_EMS01_Carrier60_Position" AT %QD10236 : DWord;
   "SDC_EMS01_Carrier61_Position" AT %QD10240 : DWord;
   "SDC_EMS01_Carrier62_Position" AT %QD10244 : DWord;
   "SDC_EMS01_Carrier63_Position" AT %QD10248 : DWord;
   "SDC_EMS01_Carrier64_Position" AT %QD10252 : DWord;
   "SDC_EMS01_Carrier65_Position" AT %QD10256 : DWord;
   "SDC_EMS01_Carrier66_Position" AT %QD10260 : DWord;
   "SDC_EMS01_Carrier67_Position" AT %QD10264 : DWord;
   "SDC_EMS01_Carrier68_Position" AT %QD10268 : DWord;
   "SDC_EMS01_Carrier69_Position" AT %QD10272 : DWord;
   "SDC_EMS01_Carrier70_Position" AT %QD10276 : DWord;
   "SDC_EMS01_Carrier71_Position" AT %QD10280 : DWord;
   "SDC_EMS01_Carrier72_Position" AT %QD10284 : DWord;
   "SDC_EMS01_Carrier73_Position" AT %QD10288 : DWord;
   "SDC_EMS01_Carrier74_Position" AT %QD10292 : DWord;
   "SDC_EMS01_Carrier75_Position" AT %QD10296 : DWord;
   "SDC_EMS01_Carrier76_Position" AT %QD10300 : DWord;
   "SDC_EMS01_Carrier77_Position" AT %QD10304 : DWord;
   "SDC_EMS01_Carrier78_Position" AT %QD10308 : DWord;
   "SDC_EMS01_Carrier79_Position" AT %QD10312 : DWord;
   "SDC_EMS01_Carrier80_Position" AT %QD10316 : DWord;
   "SDC_EMS01_Carrier81_Position" AT %QD10320 : DWord;
   "SDC_EMS01_Carrier82_Position" AT %QD10324 : DWord;
   "SDC_EMS01_Status" AT %QW11280 : Word;
   "SDC_EMS01_Faulted" AT %Q11280.1 : Bool;
   "SDC_EMS01_SpareB.2" AT %Q11280.2 : Bool;
   "SDC_EMS01_SpareB.3" AT %Q11280.3 : Bool;
   "SDC_EMS01_SpareB.4" AT %Q11280.4 : Bool;
   "SDC_EMS01_SpareB.5" AT %Q11280.5 : Bool;
   "SDC_EMS01_SpareB.6" AT %Q11280.6 : Bool;
   "SDC_EMS01_SpareB.7" AT %Q11280.7 : Bool;
   "SDC_EMS01_SpareB.8" AT %Q11281.0 : Bool;
   "SDC_EMS01_SpareB.9" AT %Q11281.1 : Bool;
   "SDC_EMS01_SpareB.10" AT %Q11281.2 : Bool;
   "SDC_EMS01_SpareB.11" AT %Q11281.3 : Bool;
   "SDC_EMS01_SpareB.12" AT %Q11281.4 : Bool;
   "SDC_EMS01_SpareB.13" AT %Q11281.5 : Bool;
   "SDC_EMS01_SpareB.14" AT %Q11281.6 : Bool;
   "SDC_EMS01_HeartBeat" AT %Q11281.7 : Bool;
   "SDC_EMS01_SpareB.16" AT %Q11282.0 : Bool;
   "SDC_EMS01_SpareB.17" AT %Q11282.1 : Bool;
   "SDC_EMS01_SpareB.18" AT %Q11282.2 : Bool;
   "SDC_EMS01_SpareB.19" AT %Q11282.3 : Bool;
   "SDC_EMS01_SpareW" AT %QW11284 : Word;
   "SDC_EMS01_FAULTS" AT %QW11286 : Word;
   "SDC_EMS01_Carrier26_Position" AT %QD10100 : DWord;
   "SDC_EMS01_Carrier27_Position" AT %QD10104 : DWord;
END_VAR

TYPE "UDT_SDCOutFaults"
VERSION : 0.1
   STRUCT
      DuplicateCarrierFault : Bool;
      MotionOnFault : Bool;
      MotionOffFault : Bool;
      CarrierSpacingFault : Bool;
   END_STRUCT;
END_TYPE

TYPE "UDT_Stop"
VERSION : 0.1
   STRUCT
      StopNumber : Bool;
      StopPosition : Bool;
      ClearToRelease : Bool;
      CarrierPresentStop : Bool;
   END_STRUCT;
END_TYPE

TYPE "UDT_HMIZonePositionStructure"
   STRUCT
      ZonePosition : Word;
      CarrierNumber : Word;
      CarrierPosition : Word;
      Faulted : Bool;
   END_STRUCT;
END_TYPE

TYPE "UDT_System"
VERSION : 0.1
   STRUCT
      Zone : Array[0..65] of "UDT_ZoneStructure";
      Carrier : Array[0..99] of "UDT_CarrierStructure";
      LowSpeedSetpoint : Word;
      HighSpeedSetpoint : Word;
      DecelPositionOffset : Word;
      SDC_Faults : Array[0..9] of Int;
      Carrier_Spacing : Int;
      TotalZones : Int;
      TotalZonePosn : Int;
      TotalCarriers : Int;
      CoarsePositionTolerance : Word;
      FinePositionTolerance : Word;
      CoarsePositionDecelOffset : Word;
      FinePositionDecelOffset : Word;
      Production_Spacing : Word;
      ClearOfStopDist : Word;
      FineDecelSpeed : Word;
      CoarseDecelSpeed : Word;
      ProductionZnSpeed : Word;
      AccumZnSpeed : Word;
      SDC : "UDT_SDC";
   END_STRUCT;
END_TYPE

TYPE "UDT_Carrier"
VERSION : 0.1
   STRUCT
      CARRIER : Array[1..99] of "UDT_CarrierStructure";
   END_STRUCT;
END_TYPE

TYPE "UDT_SDC_IN"